REGION Network 2: Error handling
         A     #IN_Reset_fault_Fkt;
         R     #Temp_IO_Fault.FLT_Motorprotection;
         R     #Temp_IO_Fault.FLT_Min_Level;
         R     #Temp_IO_Fault.FLT_WRN_C_Max;
         R     #Temp_IO_Fault.FLT_C_Max;
         R     #Temp_IO_Fault.FLT_Filter_HP;
         R     #Temp_IO_Fault.FLT_Filter_backflow;
         R     #Temp_IO_Fault.FLT_cable_break;
         R     #Temp_IO_Fault.FLT_P_Max;
   //-----
         A     #IN_MotorProtection;
         AN    #Temp_IO_Fault.FLT_Motorprotection;
         S     #Temp_IO_Fault.FLT_Motorprotection;
         S     #IO_NewFault;
   //-----
         AN    #IN_Min_Level;
         AN    #Temp_IO_Fault.FLT_Min_Level;
         S     #Temp_IO_Fault.FLT_Min_Level;
         S     #IO_NewFault;
   //-----
         A     #IN_C_OilCooling;
         A     #Temp_IO_Status.Switch_on_Motor;
         =     #Temp_IO_Status.Act_Oilcooling;
   //-----
         AN    #IN_C_Max;
         AN    #Temp_IO_Fault.FLT_WRN_C_Max;
         S     #Temp_IO_Fault.FLT_WRN_C_Max;
         S     #IO_NewFault;
   //-----
         A     #Temp_IO_Fault.FLT_WRN_C_Max;
         L     S5T#5M;
         SD    #IN_Temperatur_Timer;
         A     #IN_Temperatur_Timer;
         AN    #Temp_IO_Fault.FLT_C_Max;
         S     #Temp_IO_Fault.FLT_C_Max;
         S     #IO_NewFault;
   //-----
         A     #Temp_IO_Status.Startup_Motor_finished;
         AN    #IN_F_Filter_ReturnLine;
         L     #IN_Delay_FilterError;
         SD    #IN_Filter_Timer;
   //-----
         AN    #IN_F_Filter_FeedLine;
         AN    #Temp_IO_Fault.FLT_Filter_HP;
         S     #Temp_IO_Fault.FLT_Filter_HP;
         S     #IO_NewFault;
   //-----
         A     #IN_Filter_Timer;
         AN    #IN_F_Filter_ReturnLine;
         AN    #Temp_IO_Fault.FLT_Filter_backflow;
         S     #Temp_IO_Fault.FLT_Filter_backflow;
         S     #IO_NewFault;
   //-----
         AN    #IN_P_lowerlimit;
         AN    #IN_P_upperLimit;
         S     #Temp_IO_Fault.FLT_cable_break;
         S     #IO_NewFault;
   //-----
         O     #IN_PRequestCycle;
         ON    #Temp_IO_Status.Startup_Motor_finished;
         O     #Temp_IO_Status.Request_from_CP;
         JC    NoFP;
   //-----
         L     #IN_P_BuildUpTime;
         AN    #Temp_IO_Status.MH_Hyd_OK;
         JC    TIME;
         L     #IN_P_OperationTime;
   TIME: NOP   0;
         A     #IN_P_upperLimit;
         A     #Temp_IO_Status.Act_PressureBuildUp;
         SD    #IN_Hydraulictimer;
         A     #IN_Hydraulictimer;
         AN    #Temp_IO_Fault.FLT_P_Max;
         S     #Temp_IO_Fault.FLT_P_Max;
         S     #IO_NewFault;
   //-----
   NoFP: NOP   0;
   //-----
END_REGION

REGION Network 3: An actual fault exist
   //-----
         O     #Temp_IO_Fault.FLT_Min_Level;
         O     #Temp_IO_Fault.FLT_Motorprotection;
         O     #Temp_IO_Fault.FLT_C_Max;
         O     #Temp_IO_Fault.FLT_P_Max;
         O     #Temp_IO_Fault.FLT_cable_break;
         O     #Temp_IO_Fault.FLT_WRN_C_Max;
         O     #Temp_IO_Fault.FLT_Filter_HP;
         O     #Temp_IO_Fault.FLT_Filter_backflow;
         =     #Temp_IO_Status.Fault_Exist;
   //-----
         O     #Temp_IO_Fault.FLT_Min_Level;
         O     #Temp_IO_Fault.FLT_Motorprotection;
         O     #Temp_IO_Fault.FLT_C_Max;
         O     #Temp_IO_Fault.FLT_P_Max;
         O     #Temp_IO_Fault.FLT_cable_break;
         =     #Temp_IO_Status.FaultLevel_1;
         S     #IO_FaultLevel_1;
   //-----
         O     #Temp_IO_Fault.FLT_WRN_C_Max;
         =     #Temp_IO_Status.FaultLevel_2;
         S     #IO_FaultLevel_2;
   //-----
         O     #Temp_IO_Fault.FLT_Filter_HP;
         O     #Temp_IO_Fault.FLT_Filter_backflow;
         =     #Temp_IO_Status.FaultLevel_3;
         S     #IO_FaultLevel_3;
   //-----
END_REGION

REGION Network 4
   //-----
         L     #IN_SwitchOffTime;
         T     #Temp_Motor_ON;
   //-----
         CALL  T_CONV
         ( IN  := #Temp_Motor_ON,
           OUT := #Temp_Motor_ON_ms
         );
   //-----
         L     #Temp_Motor_ON_ms;
         L     0;
         ==I;
         =     #Temp_No_switch_OFF;
   //-----
         L     #Temp_Motor_ON_ms;
         L     60000;  // 60 sec
         <D;
         =     #Temp_DelayTimeZero;
   //-----
END_REGION

REGION Network 5
   //-----
         O     #IN_ShotStroke_by_Piston;
         ON    #IN_KK_Manager_active;
         A     #IN_PRequestCycle;
         ON    #IN_P_lowerlimit;
         O     #Temp_IO_Status.Request_from_CP;
         O     #Temp_IO_Status.Act_Oilcooling;
         A     #Temp_IO_Status.MH_Hyd_OK;
         ON    #Temp_IO_Status.MH_Hyd_OK;
         AN    #Temp_No_switch_OFF;
         AN    #Temp_DelayTimeZero;
         L     #IN_SwitchOffTime;
         SF    #IN_SwitchOFFTimer;
         A     #IN_SwitchOFFTimer;
         =     #Temp_Motor_ON_Auto;
   //-----
         AN    #IN_OPMode_Automatic;
         R     #IN_SwitchOFFTimer;
   //-----
         O     #Temp_No_switch_OFF;
         O     #Temp_DelayTimeZero;
         O     #Temp_IO_Fault.Spare14;
         S     #Temp_Motor_ON_Auto;
   //-----
END_REGION

REGION Network 6: Request hydraulic
         O     #Temp_IO_Fault.FLT_Motorprotection;
         O     #Temp_IO_Fault.FLT_Min_Level;
         O     #Temp_IO_Fault.FLT_C_Max;
         O     #Temp_IO_Fault.FLT_cable_break;
         O     #Temp_IO_Fault.FLT_P_Max;
         =     #Temp_Fault_Hyd;
   //
         AN    #IN_Pos_of_Pause_ok;
         A     #IN_KK_Manager_active;
         ON    #IN_PauseTime;
         A     #Temp_IO_Status.Switch_Hydraulic_ON_OFF;
         A     #IN_OPMode_Manual;
         O     #IN_OPMode_Automatic;
         AN    #Temp_Fault_Hyd;
         AN    #IN_Fault_from_Extern;
         =     #Temp_IO_Status.Switch_on_Motor;
   //-
         A     #Temp_Motor_ON_Auto;
         A     #IN_OPMode_Automatic;
         O     #IN_OPMode_Manual;
         A     #Temp_IO_Status.Switch_on_Motor;
         =     #Temp_Switch_Motor_ON;
END_REGION

REGION Network 7: Motor control
         A     #Temp_IO_Status.Startup_Motor_finished;
         JC    NoM;
   //
         A     #Temp_Switch_Motor_ON;
         AN    #Temp_IO_Status.Act_Star;
         AN    #IN_Hydraulictimer;
         S     #Temp_IO_Status.Act_Main;
         S     #Temp_IO_Status.Act_Star;
         L     #IN_Star_Delta_Timer;
         SE    #IN_Hydraulictimer;
   //
         A     #Temp_Switch_Motor_ON;
         A     #Temp_IO_Status.Act_Star;
         AN    #IN_Hydraulictimer;
         S     #Temp_IO_Status.Startup_Motor_finished;
         R     #IN_Hydraulictimer;
   //
         A     #Temp_IO_Status.Startup_Motor_finished;
         AN    #Temp_IO_Status.MH_Hyd_OK;
         S     #Temp_IO_Status.Act_PressureBuildUp;
   //
   NoM:  NOP   0;
         AN    #Temp_Switch_Motor_ON;
         R     #Temp_IO_Status.Startup_Motor_finished;
         R     #Temp_IO_Status.Act_Main;
         R     #Temp_IO_Status.Act_Star;
         R     #Temp_IO_Status.Act_Delta;
   //
         AN    #Temp_IO_Status.Switch_on_Motor;
         R     #Temp_IO_Status.MH_Hyd_OK;
         R     #Temp_IO_Status.Act_PressureBuildUp;
END_REGION

REGION Network 8: Pressure valve control
   // Das Druckaufbauventil für die MK- Hydraulik wird angesteuert:
   // - Nachdem die Hydaulik angefordert wird (BA Auto oder Hydraulik EIN)
   // - Bei Anforderung aus dem Zyklusbaustein (3 Sekunden vor Ende der KLZ1 und
   //   der Schuß läuft), wenn es sich um eine Kolbenmaschine handelt muß der
   //   Schußhub laufen bei einer Pumpenmaschine sofort.
   // - Bei Anforderung aus dem Reinigungsbausteinen für die dauer von x Sekunden
         AN    #IN_P_upperLimit;
         A     #Temp_IO_Status.Act_PressureBuildUp;
         S     #Temp_IO_Status.MH_Hyd_OK;
         R     #Temp_IO_Status.Act_PressureBuildUp;
   //
         O     #IN_ShotStroke_by_Piston;
         ON    #IN_KK_Manager_active;
         A     #IN_PRequestCycle;
         AN    #IN_Option2SetPoints;
         ON    #IN_P_lowerlimit;
         O     #Temp_IO_Status.Request_from_CP;
         A     #Temp_IO_Status.Startup_Motor_finished;
         A     #Temp_IO_Status.MH_Hyd_OK;
         S     #Temp_IO_Status.Act_PressureBuildUp;
   //
         A     #Temp_IO_Status.MH_Hyd_OK;
         A     #Temp_IO_Status.Request_from_CP;
         A     #Temp_IO_Status.Startup_Motor_finished;
         JCN   NoRK;
   //
         SET;
         L     #IN_P_ClPistonTime;
         SE    #IN_Hydraulictimer;
   //
         AN    #IN_Hydraulictimer;
         R     #Temp_IO_Status.Request_from_CP;
         R     #IN_Hydraulictimer;
   //
   NoRK: NOP   0;
END_REGION

REGION Network 9: Outputs
   // Die hier praktizierte Art der Ansteuerung hat den Vorteil, dass die Parameter 
   // extern mit Dummys belegt werden können, wenn sie nicht gebraucht werden.
         A     #Temp_IO_Status.Act_PressureBuildUp;
         =     #OUT_PressureValve;
         A     #Temp_IO_Status.Act_Main;
         =     #OUT_Motor_MainsContactor;
         A     #Temp_IO_Status.Act_Star;
         =     #OUT_Motor_Star;
         A     #Temp_IO_Status.Act_Delta;
         =     #OUT_Motor_Delta;
         A     #Temp_IO_Status.Act_Oilcooling;
         =     #OUT_V_OilCooling;
         A     #Temp_IO_Status.MH_Hyd_OK;
         =     #OUT_Hydraulic_active;
END_REGION

REGION Network 10: State of drive: 1-> ON; 2-> Faulty; 3->Selected but not ON
         A     #Temp_IO_Status.MH_Hyd_OK;
         L     1;
         JC    tran;
   //-
         A     #Temp_IO_Status.Fault_Exist;
         L     2;
         JC    tran;
   //-
         A     #Temp_IO_Status.Switch_Hydraulic_ON_OFF;
         AN    #Temp_IO_Status.MH_Hyd_OK;
         L     3;
         JC    tran;
   //-
         L     0;
   tran: T     #Temp_IO_Status.State_Hydraulic;
END_REGION

REGION Network 11: Save data
   //-----
         CALL  BLKMOV
         ( SRCBLK  := #Temp_IO_Status,
           RET_VAL := #ERROR_CODE,
           DSTBLK  := #Anyzeiger1
         );
   //-----
         CALL  BLKMOV
         ( SRCBLK  := #Temp_IO_Fault,
           RET_VAL := #ERROR_CODE,
           DSTBLK  := #Anyzeiger2
         );
   //-----
END_REGION
END_FUNCTION

FUNCTION "FC025_Oszilloskop" : Void   // FC25, SCL
{ S7_Optimized_Access := 'FALSE' }
VERSION : 0.1
   VAR_TEMP
      i : Int;
      Baugruppe : Int;
      Index : Int;
      Wert : Int;
      connection : Int;
   END_VAR
BEGIN
   FOR #i := 1 TO 8 DO

     CASE "DB025_Oszilloskop".Graph[#i].Auswahl OF
       10:  CASE "DB025_Oszilloskop".Graph[#i].Komponente OF // Adresse
             20:  CASE "DB025_Oszilloskop".Graph[#i].Sensor OF  // Datenbaustein
                 101: "DB025_Oszilloskop".Graph[#i].Wert :=        // Bool
                     INT_TO_REAL(BOOL_TO_INT( PEEK_BOOL(area:=16#84,dbNumber:=WORD_TO_UINT("DB025_Oszilloskop".Graph[#i].DB_Nummer),byteOffset:="DB025_Oszilloskop".Graph[#i].Adresse,bitOffset:="DB025_Oszilloskop".Graph[#i].Bit) ) ) * "DB025_Oszilloskop".Graph[#i].Skalierung;  
                 102: "DB025_Oszilloskop".Graph[#i].Wert :=        // Byte
                     INT_TO_REAL( PEEK_BYTE(area:=16#84,dbNumber:=WORD_TO_UINT("DB025_Oszilloskop".Graph[#i].DB_Nummer),byteOffset:="DB025_Oszilloskop".Graph[#i].Adresse) ) * "DB025_Oszilloskop".Graph[#i].Skalierung; 
                 103: "DB025_Oszilloskop".Graph[#i].Wert :=        // Int
                     INT_TO_REAL( PEEK_WORD(area:=16#84,dbNumber:=WORD_TO_UINT("DB025_Oszilloskop".Graph[#i].DB_Nummer),byteOffset:="DB025_Oszilloskop".Graph[#i].Adresse) ) * "DB025_Oszilloskop".Graph[#i].Skalierung; 
                 104: "DB025_Oszilloskop".Graph[#i].Wert :=        // Dint
                     DINT_TO_REAL( PEEK_DWORD(area:=16#84,dbNumber:=WORD_TO_UINT("DB025_Oszilloskop".Graph[#i].DB_Nummer),byteOffset:="DB025_Oszilloskop".Graph[#i].Adresse) ) * "DB025_Oszilloskop".Graph[#i].Skalierung; 
                 105: "DB025_Oszilloskop".Graph[#i].Wert :=        // Real
                     DINT_TO_REAL( PEEK_DWORD(area:=16#84,dbNumber:=WORD_TO_UINT("DB025_Oszilloskop".Graph[#i].DB_Nummer),byteOffset:="DB025_Oszilloskop".Graph[#i].Adresse) ) * "DB025_Oszilloskop".Graph[#i].Skalierung; 
                 106: "DB025_Oszilloskop".Graph[#i].Wert :=        // Timer
                     REAL#0.0; 
               ELSE
                 "DB025_Oszilloskop".Graph[#i].Wert :=  REAL#0.0;
               END_CASE;
             21:  CASE "DB025_Oszilloskop".Graph[#i].Sensor OF  // Eingang
                 101: "DB025_Oszilloskop".Graph[#i].Wert :=        // Bool
                     INT_TO_REAL(BOOL_TO_INT( PEEK_BOOL(area:=16#81,dbNumber:=0,byteOffset:="DB025_Oszilloskop".Graph[#i].Adresse,bitOffset:="DB025_Oszilloskop".Graph[#i].Bit) ) ) * "DB025_Oszilloskop".Graph[#i].Skalierung;
                 102: "DB025_Oszilloskop".Graph[#i].Wert :=        // Byte
                     INT_TO_REAL( PEEK_BYTE(area:=16#81,dbNumber:=0,byteOffset:="DB025_Oszilloskop".Graph[#i].Adresse) ) * "DB025_Oszilloskop".Graph[#i].Skalierung; 
                 103: "DB025_Oszilloskop".Graph[#i].Wert :=        // Int
                     INT_TO_REAL( PEEK_WORD(area:=16#81,dbNumber:=0,byteOffset:="DB025_Oszilloskop".Graph[#i].Adresse) ) * "DB025_Oszilloskop".Graph[#i].Skalierung; 
                 104: "DB025_Oszilloskop".Graph[#i].Wert :=        // Dint
                     DINT_TO_REAL( PEEK_DWORD(area:=16#81,dbNumber:=0,byteOffset:="DB025_Oszilloskop".Graph[#i].Adresse) ) * "DB025_Oszilloskop".Graph[#i].Skalierung; 
                 105: "DB025_Oszilloskop".Graph[#i].Wert :=        // Real
                     REAL#0.0 ; 
               ELSE
                 "DB025_Oszilloskop".Graph[#i].Wert :=  REAL#0.0;
               END_CASE;
             22:  CASE "DB025_Oszilloskop".Graph[#i].Sensor OF  // Ausgang
                 101: "DB025_Oszilloskop".Graph[#i].Wert :=        // Bool
                     INT_TO_REAL(BOOL_TO_INT( PEEK_BOOL(area:=16#82,dbNumber:=0,byteOffset:="DB025_Oszilloskop".Graph[#i].Adresse,bitOffset:="DB025_Oszilloskop".Graph[#i].Bit) ) ) * "DB025_Oszilloskop".Graph[#i].Skalierung;
                 102: "DB025_Oszilloskop".Graph[#i].Wert :=        // Byte
                     INT_TO_REAL( PEEK_BYTE(area:=16#82,dbNumber:=0,byteOffset:="DB025_Oszilloskop".Graph[#i].Adresse) ) * "DB025_Oszilloskop".Graph[#i].Skalierung; 
                 103: "DB025_Oszilloskop".Graph[#i].Wert :=        // Int
                     INT_TO_REAL( PEEK_WORD(area:=16#82,dbNumber:=0,byteOffset:="DB025_Oszilloskop".Graph[#i].Adresse) ) * "DB025_Oszilloskop".Graph[#i].Skalierung; 
                 104: "DB025_Oszilloskop".Graph[#i].Wert :=        // Dint
                     DINT_TO_REAL( PEEK_DWORD(area:=16#82,dbNumber:=0,byteOffset:="DB025_Oszilloskop".Graph[#i].Adresse) ) * "DB025_Oszilloskop".Graph[#i].Skalierung; 
                 105: "DB025_Oszilloskop".Graph[#i].Wert :=        // Real
                     DINT_TO_REAL( PEEK_DWORD(area:=16#82,dbNumber:=0,byteOffset:="DB025_Oszilloskop".Graph[#i].Adresse) ) * "DB025_Oszilloskop".Graph[#i].Skalierung; 
               ELSE
                 "DB025_Oszilloskop".Graph[#i].Wert :=  REAL#0.0;
               END_CASE;
             23:  CASE "DB025_Oszilloskop".Graph[#i].Sensor OF  // Merker
                 101: "DB025_Oszilloskop".Graph[#i].Wert :=       // Bool
                     INT_TO_REAL(BOOL_TO_INT( PEEK_BOOL(area:=16#83,dbNumber:=0,byteOffset:="DB025_Oszilloskop".Graph[#i].Adresse,bitOffset:="DB025_Oszilloskop".Graph[#i].Bit) ) ) * "DB025_Oszilloskop".Graph[#i].Skalierung;
                 102: "DB025_Oszilloskop".Graph[#i].Wert :=        // Byte
                     INT_TO_REAL( PEEK_BYTE(area:=16#83,dbNumber:=0,byteOffset:="DB025_Oszilloskop".Graph[#i].Adresse) ) * "DB025_Oszilloskop".Graph[#i].Skalierung; 
                 103: "DB025_Oszilloskop".Graph[#i].Wert :=        // Int
                     INT_TO_REAL( PEEK_WORD(area:=16#83,dbNumber:=0,byteOffset:="DB025_Oszilloskop".Graph[#i].Adresse) ) * "DB025_Oszilloskop".Graph[#i].Skalierung; 
                 104: "DB025_Oszilloskop".Graph[#i].Wert :=        // Dint
                     DINT_TO_REAL( PEEK_DWORD(area:=16#83,dbNumber:=0,byteOffset:="DB025_Oszilloskop".Graph[#i].Adresse) ) * "DB025_Oszilloskop".Graph[#i].Skalierung; 
                 105: "DB025_Oszilloskop".Graph[#i].Wert :=         // Real
                     DINT_TO_REAL( PEEK_DWORD(area:=16#83,dbNumber:=0,byteOffset:="DB025_Oszilloskop".Graph[#i].Adresse) ) * "DB025_Oszilloskop".Graph[#i].Skalierung; ; 
               ELSE
                 "DB025_Oszilloskop".Graph[#i].Wert :=  REAL#0.0;
               END_CASE;
             24:  CASE "DB025_Oszilloskop".Graph[#i].Sensor OF  // Timer
                 106: "DB025_Oszilloskop".Graph[#i].Wert := REAL#0.0 ; // Timer
               ELSE
                 "DB025_Oszilloskop".Graph[#i].Wert :=  REAL#0.0;
               END_CASE;
           ELSE
             "DB025_Oszilloskop".Graph[#i].Wert :=  REAL#0.0;
           END_CASE;
       40:  CASE "DB025_Oszilloskop".Graph[#i].Sensor OF       // Behälter
             1:  "DB025_Oszilloskop".Graph[#i].Wert :=         // Durchfluss
                 REAL#0.0;               
             2:  "DB025_Oszilloskop".Graph[#i].Wert :=         // Druck
                 "DB602_PV_Tank".Tank["DB025_Oszilloskop".Graph[#i].Komponente].Pressure.PV_ActV.Value   * "DB025_Oszilloskop".Graph[#i].Skalierung;    
             3:  "DB025_Oszilloskop".Graph[#i].Wert :=         // Füllstand
                 "DB602_PV_Tank".Tank["DB025_Oszilloskop".Graph[#i].Komponente].Level.PV_ActV.Value      * "DB025_Oszilloskop".Graph[#i].Skalierung;         
             4:  "DB025_Oszilloskop".Graph[#i].Wert :=         // Gasbeladung
                 "DB602_PV_Tank".Tank["DB025_Oszilloskop".Graph[#i].Komponente].Nucleation.PV_ActV.Value * "DB025_Oszilloskop".Graph[#i].Skalierung;  
             5:  "DB025_Oszilloskop".Graph[#i].Wert :=         // Mischungsverhältnis         
                 REAL#40.0;              
             6:  "DB025_Oszilloskop".Graph[#i].Wert :=         // Temperatur
                 "DB602_PV_Tank".Tank["DB025_Oszilloskop".Graph[#i].Komponente].Temp.PV_ActV.Value       * "DB025_Oszilloskop".Graph[#i].Skalierung;        
           ELSE
             "DB025_Oszilloskop".Graph[#i].Wert :=  REAL#0.0;
           END_CASE;
        30:  CASE "DB025_Oszilloskop".Graph[#i].Sensor OF      // Pumpe
             1:  "DB025_Oszilloskop".Graph[#i].Wert :=         // Durchfluss
                 "DB608_PV_Metering".Metering["DB025_Oszilloskop".Graph[#i].Komponente].Flow.PV_ActV.Value *"DB025_Oszilloskop".Graph[#i].Skalierung;       
             2:  "DB025_Oszilloskop".Graph[#i].Wert :=         // Druck
                 "DB608_PV_Metering".Metering["DB025_Oszilloskop".Graph[#i].Komponente].Pressure.PV_ActV.Value  * "DB025_Oszilloskop".Graph[#i].Skalierung;    
             3:  "DB025_Oszilloskop".Graph[#i].Wert :=         // Füllstand
                 REAL#0.0;   
             4:  "DB025_Oszilloskop".Graph[#i].Wert :=         // Gasbeladung
                 REAL#0.0; 
             5:  "DB025_Oszilloskop".Graph[#i].Wert :=         // Mischungsverhältnis
                 "DB608_PV_Metering".Metering["DB025_Oszilloskop".Graph[#i].Komponente].MixingRatio.PV_ActV.Value  * "DB025_Oszilloskop".Graph[#i].Skalierung; 
             6:  "DB025_Oszilloskop".Graph[#i].Wert :=         // Temperatur
                 "DB608_PV_Metering".Metering["DB025_Oszilloskop".Graph[#i].Komponente].Temperature.PV_ActV.Value  * "DB025_Oszilloskop".Graph[#i].Skalierung; 
           ELSE
             "DB025_Oszilloskop".Graph[#i].Wert :=  REAL#0.0;
           END_CASE;
        20: #connection := 0;
                IF "DB025_Oszilloskop".Graph[#i].Komponente = "DB704_MH_Value".Mixinghead["DB025_Oszilloskop".Graph[#i].Nummer].MH_Connection[1].Pump_No THEN #connection := 1;  
                ELSIF "DB025_Oszilloskop".Graph[#i].Komponente = "DB704_MH_Value".Mixinghead["DB025_Oszilloskop".Graph[#i].Nummer].MH_Connection[2].Pump_No THEN #connection := 2;  
                ELSIF "DB025_Oszilloskop".Graph[#i].Komponente = "DB704_MH_Value".Mixinghead["DB025_Oszilloskop".Graph[#i].Nummer].MH_Connection[3].Pump_No THEN #connection := 3;  
                ELSIF "DB025_Oszilloskop".Graph[#i].Komponente = "DB704_MH_Value".Mixinghead["DB025_Oszilloskop".Graph[#i].Nummer].MH_Connection[4].Pump_No THEN #connection := 4;  
                ELSIF "DB025_Oszilloskop".Graph[#i].Komponente = "DB704_MH_Value".Mixinghead["DB025_Oszilloskop".Graph[#i].Nummer].MH_Connection[5].Pump_No THEN #connection := 5;  
                ELSIF "DB025_Oszilloskop".Graph[#i].Komponente = "DB704_MH_Value".Mixinghead["DB025_Oszilloskop".Graph[#i].Nummer].MH_Connection[6].Pump_No THEN #connection := 6;
                ELSE #connection := 0;
                END_IF;

           CASE "DB025_Oszilloskop".Graph[#i].Sensor OF        // Mischkopf    
             1:  "DB025_Oszilloskop".Graph[#i].Wert :=         // Durchfluss
                 REAL#0.0;             
             2:  "DB025_Oszilloskop".Graph[#i].Wert :=         // Druck
                 "DB604_PV_Mixinghead".Mixinghead["DB025_Oszilloskop".Graph[#i].Nummer].Pressure_Connection[#connection].PV_ActV.Value * "DB025_Oszilloskop".Graph[#i].Skalierung;  
             3:  "DB025_Oszilloskop".Graph[#i].Wert :=         // Füllstand
                 REAL#0.0;               
             4:  "DB025_Oszilloskop".Graph[#i].Wert :=         // Gasbeladung
                 REAL#0.0;             
             5:  "DB025_Oszilloskop".Graph[#i].Wert :=         // Mischungsverhältnis
                 REAL#0.0;                     
             6:  "DB025_Oszilloskop".Graph[#i].Wert :=         // Temperatur
                 "DB604_PV_Mixinghead".Mixinghead["DB025_Oszilloskop".Graph[#i].Nummer].Temperature_Connection[#connection].PV_ActV.Value * "DB025_Oszilloskop".Graph[#i].Skalierung;    
           ELSE
             "DB025_Oszilloskop".Graph[#i].Wert :=  REAL#0.0;
           END_CASE;
     ELSE
       "DB025_Oszilloskop".Graph[#i].Wert :=  REAL#0.0;
     END_CASE;
   END_FOR;
END_FUNCTION

FUNCTION "FC041_SwitchOverUnit" : Void   // FC41, STL
TITLE = Control of switch over units
{ S7_Optimized_Access := 'FALSE' }
AUTHOR : KT242
FAMILY : RS_KK
NAME : SWU
VERSION : 1.3
   VAR_INPUT
      IN_select_piston : Bool;   // Differentiation if programmblock is used by pump- or piston metering
      IN_filling_piston : Bool;   // Component piston in filling mode, used to switchover after strokes
      IN_OperationMode_valid : Bool;   // Operation mode valid
      IN_AcknoldgeFaults : Bool;   // Quit faults
      IN_cycle_running : Bool;   // During cycle is running no. of SWO is set by foaming program
      IN_PistonService : Bool;   // Piston service is selected to activate a switch over unit
      IN_Circulation_active : Bool;   // During active recirculation SWU will be switched over after a setted time
      IN_Circulation_HP_active : Bool;   // At high pressure circulation mixinghead no. is set by selected mixinghead
      IN_MH_No_at_FoamingCycle : Byte;   // Mixinghead number from foaming program to select SWU
      IN_MH_No_at_HP_Cycle : DWord;   // Mixinghead number from program block "operation mode" to select SWU by HP
      IN_StokeCounter : Counter;   // Counter of piston strokes to switch over to MH at piston machine
      IN_Amount_Strokes : Int;   // Setting of piston strokes to switch over to MH at piston machine
      IN_FlushingTimer : Timer;   // Timer flushing components between the mixingheads
      IN_SWU_FlushingTime : S5Time;   // Flushing time at each mixinghead at recirculation -> switchover to next MH
      IN_SwitchOverTimer : Timer;   // Timer to switch off and over between SWU's -> two SWU selected
      IN_SwitchOffTime : S5Time;   // Timevalue of increased activation of SWU at switch off
      IN_SwitchOverTime : S5Time;   // Timevalue of common activation of two SWU's during switch over
   END_VAR
   VAR_IN_OUT
      IO_Status : ANY;   // Speichern der Umschalteinheiten (USE)- Zustände für das Programm
      IO_Fault : ANY;
      IO_NewFault : Bool;
      IO_FaultLevel_1 : Bool;
      IO_FaultLevel_2 : Bool;
      IO_FaultLevel_3 : Bool;
   END_VAR
   VAR_TEMP
      Temp_IO_Status : "UDT041_SWU_State";
      TEMP_IO_Fault : "UDT1841_FLT_SWU";
      ERROR_CODE : Int;   // Error state of systemfunction "BLKMOV" Blockmove
      Anyzeiger1 : ANY;   // Pointer to copy thr array "IO_Status" and "Temp_IO_Status"
      Anyzeiger2 : ANY;   // Pointer to copy thr array "IO_Status" and "Temp_IO_Status"
      Baustein_Nr : Int;   // Merker zur Erkennung des Speicherbereiches der Bits "IO_Ziel_USE"
      Adresse_im_Baustein : DWord;   // and the start adress within the program block
      Freigaben_lokal : DWord;   // Intermidiate flags of release of switch over units (from UDT to DWORD)
      USE_Ventile_lokal : DWord;   // Zwischenspeicher der angesteuerten Umschalteinheiten (von UDT auf DWORD)
      Angef_USE_Nummer_lokal : DWord;   // Zwischenspeicher der angeforderten Umschalteinheiten (von UDT auf DWORD)
      Ziel_USE_lokal : DWord;   // Zwischenspeicher der auzusteuernden Umschalteinheiten (von UDT auf DWORD)
      U_A_Zeitwert : S5Time;   // Zeitwert bei der Unterscheidung ob eine USE um- oder abgeschaltet werden soll
      Temp_SWU_FlushingTime : S5Time;   // Zeitwert für die Spülzeit mindestens 3 Sekunden
      Spuelzeit_laeuft : Bool;   // Die Spülzeit der einzelnen Mischköpfe (USE) läuft und wird durchgetaktet
      Abschaltzeit_laeuft : Bool;   // Die Abschaltzeit der offenen USE läuft -> keine weitere USE angefordert
      Wiedereinschaltung : Bool;   // Es wurde innerhalb der Abschaltzeit Kreislauf etc. angeschaltet
   END_VAR
BEGIN

REGION Network 1: Saved data integration
   // Änderungen:
   // -------------------------------------------------------------------------------
   // Durch die Verwendung von + -1 bei der Ermittlung der angeforderten USE während 
   // des Zyklusses (Netzwerk 5) sind nur bis zu 16 Mischköpfe ansteuerbar.
   // Durch das umsetzen in Doppelworte (L     DW#16#1) wird eine Ansteuerung bis zu 
   // 32 Mischköpfe möglich
   // 
   // v.d.Geest       19.01.2005
   // -------------------------------------------------------------------------------
   // Wenn im Rechner ein Mischkopf als folgender Teilschuß angewählt wurde, dessen 
   // USE aber nicht freigegeben war kam es zu einer Max. Druck- Störung.
   // Um dieses zu vermeiden wurde eine neue Störung "USE_nicht_freigegeben" im 
   // Netzwerk 7 ab Zeile 49 eingebunden.
   // 
   // v.d.Geest       27.10.2003
   // -------------------------------------------------------------------------------
   // Die Ansteuerung der "Um_Abschaltzeit" funktionierte so nicht:
   // Bei Anwahl Kreislauf aus dem Stillstand lief die "Um_Abschaltzeit" ab, obwohl 
   // vorher kein weiterer Mischkopf angewählt wurde. 
   // Ebenso wurde die gesamte Abschaltzeit abgewartet wenn zwischen dem Auschalten 
   // des Kreislaufes über zB. MK01 und dem winschalten des Kreislaufes über zB. MK02 
   // weniger als 5 Sekunden (Abschaltzeit) lagen.
   // Die Auswirkungen waren zu spüren der Anwahl des HD- Kreislaufes, da dieser erst 
   // gestartet wurde wenn die "Um_Abschaltzeit" abgelaufen war.
   // Das alte Bit "Um_Abschaltzeit" im UDT wurde in "Umschaltzeit" (wichtig bei 
   // schnellem Druckaufbau und bei Ansteuerung des Reinigungskolbens) umbenannt und 
   // ein neues Bit "Abschaltzeit" wurde erstellt.
   // Bei Übernahme bitte UDT 41 mit einspielen.
   // 
   // v.d.Geest       11.04.2003
   // -------------------------------------------------------------------------------
         LAR1;
         L;
         LAR2;
   //
         L     W[AR2, P#0.0];  // Bytes
         T     W[AR1, P#0.0];
         L     W [ AR2 , P#2.0 ];  // Amount of bytes
         T     W[AR1, P#2.0];
         L     W [ AR2 , P#4.0 ];  // Block no,
         T     W[AR1, P#4.0];
         L     D [ AR2 , P#6.0 ];  // Startadress of datas
         T     D[AR1, P#6.0];
   //
         CALL  BLKMOV
         ( SRCBLK  := #Anyzeiger1,
           RET_VAL := #ERROR_CODE,
           DSTBLK  := #Temp_IO_Status
         );

         LAR1;
         L;
         LAR2;
   //
         L     W[AR2, P#0.0];  // Bytes
         T     W[AR1, P#0.0];
         L     W [ AR2 , P#2.0 ];  // Amount of bytes
         T     W[AR1, P#2.0];
         L     W [ AR2 , P#4.0 ];  // Block no,
         T     W[AR1, P#4.0];
         L     D [ AR2 , P#6.0 ];  // Startadress of datas
         T     D[AR1, P#6.0];
   //
         CALL  BLKMOV
         ( SRCBLK  := #Anyzeiger2,
           RET_VAL := #ERROR_CODE,
           DSTBLK  := #TEMP_IO_Fault
         );
   //
END_REGION

REGION Network 2: Störungen quittieren
         A     #IN_AcknoldgeFaults;
         R     #TEMP_IO_Fault.FLT_open_SWU_disabelt;
         R     #TEMP_IO_Fault.FLT_No_SWU_selected;
         R     #TEMP_IO_Fault.FLT_Sel_SWU_not_released;
END_REGION

REGION Network 3: Datenschieben
   //_______________________________________________________________
   // Schieben der USE- Freigaben auf lokalen DWord- Bereich
   //
         L;
         LAR2;
         L;
         LAR1;
   //
         L     LD [ AR2 , P#8.0 ];
         T     LD[AR1, P#0.0];
   //_______________________________________________________________
   // Schieben der Ziel- USE vom Rechner auf lokalen DWord- Bereich
   //
         L;
         LAR2;
         L;
         LAR1;
   //
         L     LD [ AR2 , P#12.0 ];
         T     LD[AR1, P#0.0];
   //_______________________________________________________________
   // Schieben der offenen USE auf lokalen DWord- Bereich
   //
         L;
         LAR1;
   //
         L     LD [ AR2 , P#16.0 ];
         T     LD[AR1, P#0.0];
END_REGION

REGION Network 4: Allgemein Verwaltung der angeforderten USE
         L     #Freigaben_lokal;
         L     0;
         <>D;
         =     #Temp_IO_Status.Min_1_SWU_release;
   //
         L     #USE_Ventile_lokal;
         L     #Freigaben_lokal;
         AD;
         <>D;
         =     #Temp_IO_Status.Open_SWU_disabelt;
   //
         ON    #IN_cycle_running;
         R     #Temp_IO_Status.CycleStarted;
   //
         A     #IN_cycle_running;
         A(;
         L     #IN_MH_No_at_FoamingCycle;
         L     0;
         <>I;
         );
         O     #Temp_IO_Status.CycleStarted;
         JC    ZYKL;
   //
         A     #IN_Circulation_HP_active;
         JC    HD;
   //
         O     #IN_Circulation_active;
         O     #IN_PistonService;
         A     #Temp_IO_Status.Min_1_SWU_release;
         JC    KK;
END_REGION

REGION Network 5: Keine USE angefordert
         L     0;
         T     #Angef_USE_Nummer_lokal;
   //
         SET;
         R     #IN_StokeCounter;
         R     #Temp_IO_Status.Hubcounter_OK;
         R     #IN_FlushingTimer;
   //
         CLR;
         SP    #IN_FlushingTimer;
   //
         JU    N05A;
END_REGION

REGION Network 6: Zyklus läuft oder Kreislauf Hochdruck
   ZYKL: NOP   0;
         S     #Temp_IO_Status.CycleStarted;
   //-
         L     0;
         L     #IN_MH_No_at_FoamingCycle;
         ==I;
         JC    NoUS;
         L     16#0000_0001;
         -D;
         L     16#0000_0001;
         SLD;
         JU    Next;
   NoUS: L     #Ziel_USE_lokal;
   Next: T     #Angef_USE_Nummer_lokal;
         JU    N05A;
   //
   HD:   L     #IN_MH_No_at_HP_Cycle;
         T     #Angef_USE_Nummer_lokal;
         JU    N05A;
END_REGION

REGION Network 7: Unterscheidung RS oder KK für USE- Spülung
   KK:   AN    #IN_select_piston;
         JC    RS;
   //
         A     #IN_Circulation_active;
         A     #IN_filling_piston;
         CU    #IN_StokeCounter;
   //
         L     #IN_Amount_Strokes;
         LC    #IN_StokeCounter;
         ==I;
         R     #IN_StokeCounter;
         =     #Temp_IO_Status.Hubcounter_OK;
   //
   RS:   L     0;
         L     #Temp_IO_Status.SWU_for_Circulation;
         ==D;
         JC    ERST;
         JU    SPUE;
   ERST: L     1;
         T     #Temp_IO_Status.SWU_for_Circulation;
   //
   SPUE: L     #IN_SWU_FlushingTime;
         T     #Temp_SWU_FlushingTime;
         L     S5T#3S;
         >D;
         JC    STRT;
         T     #Temp_SWU_FlushingTime;
   //
   STRT: A(;
         AN    #IN_FlushingTimer;
         AN    #IN_select_piston;
         O;
         AN    #Temp_IO_Status.Hubcounter_OK;
         A     #IN_select_piston;
         );
         A(;
         L     #Temp_IO_Status.SWU_for_Circulation;
         L     #Freigaben_lokal;
         AD;
         ==D;
         );
         =     #Spuelzeit_laeuft;
   //
         A     #Spuelzeit_laeuft;
         AN    #IN_select_piston;
         L     #Temp_SWU_FlushingTime;
         SD    #IN_FlushingTimer;
   //
         A     #Spuelzeit_laeuft;
         JC    RED;
   //
   TAKT: L     #Temp_IO_Status.SWU_for_Circulation;
         SLD   1;
         JP    USE1;
         JU    TEST;
   //
   USE1: L     1;
   //
   TEST: T     #Temp_IO_Status.SWU_for_Circulation;
         L     #Freigaben_lokal;
         AD;
         <>D;
         JC    TAKT;
   //
   RED:  L     #Temp_IO_Status.SWU_for_Circulation;
         T     #Angef_USE_Nummer_lokal;
END_REGION

REGION Network 8: Abschaltzeit / Umschaltzeit / USE- Ansteuerung
   N05A: L     #Angef_USE_Nummer_lokal;
         L     0;
         ==D;
         =     #Abschaltzeit_laeuft;
         S     #Temp_IO_Status.Stoptime_runs;
   //
         AN    #Abschaltzeit_laeuft;
         A     #Temp_IO_Status.Stoptime_runs;
         =     #Wiedereinschaltung;
         R     #Temp_IO_Status.Stoptime_runs;
         JC    Cl_T;
   //
         L     #IN_SwitchOverTime;
         AN    #Abschaltzeit_laeuft;
         JC    Zeit;
         L     #IN_SwitchOffTime;
   Zeit: T     #U_A_Zeitwert;
   //
         A(;
         L     #Ziel_USE_lokal;  // USE_Ventile
         L     0;
         <>D;
         );
         A(;
         L     #Angef_USE_Nummer_lokal;
         L     #Ziel_USE_lokal;  // USE_Ventile
         <>D;
         );
         L     #U_A_Zeitwert;
         SE    #IN_SwitchOverTimer;
   //
         AN    #IN_SwitchOverTimer;
         R     #Temp_IO_Status.Stoptime_runs;
   //
         A     #IN_SwitchOverTimer;
         AN    #Temp_IO_Status.Stoptime_runs;
         =     #Temp_IO_Status.Switchingtime_runs;
         JU    ZUSE;
   //
   Cl_T: NOP   0;
         CLR;
         SP    #IN_SwitchOverTimer;
   //
   ZUSE: L     #Angef_USE_Nummer_lokal;
         L     #Freigaben_lokal;
         AD;
         T     #Ziel_USE_lokal;  // USE_Ventile
   //
         A(;
         L     #Angef_USE_Nummer_lokal;
         L     0;
         <>D;
         );
         A(;
         L     #Ziel_USE_lokal;  // USE_Ventile
         L     0;
         ==D;
         );
         =     #Temp_IO_Status.SWU_not_released;
   //_______________________________________________________________
   // Schieben der allein offenen USE auf den Status - Bereich
   //
         L;
         LAR2;
         L;  // USE_Ventile
         LAR1;
   //
         L     LD[AR1, P#0.0];  // USE_Ventile
         T     LD [ AR2 , P#20.0 ];  // Temp_Status.Offene_USE_allein
   //
         O     #Temp_IO_Status.Switchingtime_runs;
         O     #Temp_IO_Status.Stoptime_runs;
         JCN   OUSE;
   //
         L     #Ziel_USE_lokal;
         L     #USE_Ventile_lokal;
         OW;
         T     #USE_Ventile_lokal;
   //_______________________________________________________________
   // Ablöschen der allein offenen USE auf den Status - Bereich
   //
         L;
         LAR2;
   //
         L     0;
         T     LD [ AR2 , P#20.0 ];  // Temp_Status.Offene_USE_allein
   //
         JU    M017;
   //
   OUSE: NOP   0;
   //
         L     #Ziel_USE_lokal;
         T     #USE_Ventile_lokal;
   //
   M017: NOP   0;
   //
         L     #USE_Ventile_lokal;
         L     0;
         ==D;
         R     #Temp_IO_Status.SWU_OK;
         JC    NUSE;
   //
   M012: NOP   0;
         TAK;
         SRD   1;
         JZ    M012;
         ==I;
         =     #Temp_IO_Status.SWU_OK;
   //
   NUSE: NOP   0;
END_REGION

REGION Network 9
   //_______________________________________________________________
   // Schieben der offenen USE auf den "IO_Status"- Bereich
   //
         L;
         LAR2;
         L;
         LAR1;
   //
         L     LD[AR1, P#0.0];  // USE_Ventile
         T     LD [ AR2 , P#16.0 ];  // Temp_Status.Open_SWU
   //_______________________________________________________________
   // Schieben der lokalen Ziel- USE auf den Ziel- USE- Bereich
   //
         L;
         LAR2;
         L;
         LAR1;
         L     LD [ AR1 , P#0.0 ];  // Ziel_USE_Lokal
         T     LD [ AR2 , P#12.0 ];  // Temp_Status.Target_SWU
   //_______________________________________________________________
   //
END_REGION

REGION Network 10
         L     0;
         A     #Temp_IO_Status.Target_SWU."01";
         JCN   nMH01;
         +     1;
         JU    NoHMopen;
   nMH01:NOP   0;
         A     #Temp_IO_Status.Target_SWU."02";
         JCN   nMH02;
         +     2;
         JU    NoHMopen;
   nMH02:NOP   0;
         A     #Temp_IO_Status.Target_SWU."03";
         JCN   nMH03;
         +     3;
         JU    NoHMopen;
   nMH03:NOP   0;
         A     #Temp_IO_Status.Target_SWU."04";
         JCN   nMH04;
         +     4;
         JU    NoHMopen;
   nMH04:NOP   0;
         A     #Temp_IO_Status.Target_SWU."05";
         JCN   nMH05;
         +     5;
         JU    NoHMopen;
   nMH05:NOP   0;
         A     #Temp_IO_Status.Target_SWU."06";
         JCN   nMH06;
         +     6;
         JU    NoHMopen;
   nMH06:NOP   0;
         A     #Temp_IO_Status.Target_SWU."07";
         JCN   nMH07;
         +     7;
         JU    NoHMopen;
   nMH07:NOP   0;
         A     #Temp_IO_Status.Target_SWU."08";
         JCN   nMH08;
         +     8;
         JU    NoHMopen;
   nMH08:NOP   0;
         A     #Temp_IO_Status.Target_SWU."09";
         JCN   nMH09;
         +     9;
         JU    NoHMopen;
   nMH09:NOP   0;
         A     #Temp_IO_Status.Target_SWU."10";
         JCN   nMH10;
         +     10;
         JU    NoHMopen;
   nMH10:NOP   0;
         A     #Temp_IO_Status.Target_SWU."11";
         JCN   nMH11;
         +     11;
         JU    NoHMopen;
   nMH11:NOP   0;
         A     #Temp_IO_Status.Target_SWU."12";
         JCN   nMH12;
         +     12;
         JU    NoHMopen;
   nMH12:NOP   0;
         A     #Temp_IO_Status.Target_SWU."13";
         JCN   nMH13;
         +     13;
         JU    NoHMopen;
   nMH13:NOP   0;
         A     #Temp_IO_Status.Target_SWU."14";
         JCN   nMH14;
         +     14;
         JU    NoHMopen;
   nMH14:NOP   0;
         A     #Temp_IO_Status.Target_SWU."15";
         JCN   nMH15;
         +     15;
         JU    NoHMopen;
   nMH15:NOP   0;
         A     #Temp_IO_Status.Target_SWU."16";
         JCN   nMH16;
         +     16;
         JU    NoHMopen;
   nMH16:NOP   0;

   NoHMopen:NOP   0;
         T     #Temp_IO_Status.ActualSWU;
END_REGION

REGION Network 11: Error handling
         A     #Temp_IO_Status.Open_SWU_disabelt;
         AN    #TEMP_IO_Fault.FLT_open_SWU_disabelt;
         S     #TEMP_IO_Fault.FLT_open_SWU_disabelt;
         S     #IO_NewFault;
   //-----
         AN    #Temp_IO_Status.Min_1_SWU_release;
         A     #IN_OperationMode_valid;
         AN    #TEMP_IO_Fault.FLT_No_SWU_selected;
         S     #TEMP_IO_Fault.FLT_No_SWU_selected;
         S     #IO_NewFault;
   //-----
         A     #Temp_IO_Status.SWU_not_released;
         AN    #TEMP_IO_Fault.FLT_Sel_SWU_not_released;
         S     #TEMP_IO_Fault.FLT_Sel_SWU_not_released;
         S     #IO_NewFault;
   //-----
         O     #TEMP_IO_Fault.FLT_open_SWU_disabelt;
         O     #TEMP_IO_Fault.FLT_No_SWU_selected;
         O     #TEMP_IO_Fault.FLT_Sel_SWU_not_released;
         =     #Temp_IO_Status.FaultLevel_1;
         S     #IO_FaultLevel_1;
   //-----
         CLR;
         =     #Temp_IO_Status.FaultLevel_2;
         S     #IO_FaultLevel_2;
   //-----
         CLR;
         =     #Temp_IO_Status.FaultLevel_3;
         S     #IO_FaultLevel_3;
END_REGION

REGION Network 12: Save data
         CALL  BLKMOV
         ( SRCBLK  := #Temp_IO_Status,
           RET_VAL := #ERROR_CODE,
           DSTBLK  := #Anyzeiger1
         );
   //
         CALL  BLKMOV
         ( SRCBLK  := #TEMP_IO_Fault,
           RET_VAL := #ERROR_CODE,
           DSTBLK  := #Anyzeiger2
         );
   //
END_REGION
END_FUNCTION

FUNCTION "FC042_MixingHead" : Void   // FC42, STL
TITLE = Control of mixinghead valve
{ S7_Optimized_Access := 'FALSE' }
AUTHOR : KT242
FAMILY : RS_KK
NAME : MHead
VERSION : 1.1
   VAR_INPUT
      IN_SWU_openValve : "UDT001_DWord_1_32";
      IN_OPMode_Automatic : Bool;
      IN_OPMode_Production : Bool;
      IN_OPMode_Test : Bool;
      IN_Error_Level_1 : Bool;
      IN_SWU_OK : Bool;
      IN_Release_Foamingcycle : Bool;
      IN_ExternalRel_Foaming : Bool;
      IN_ToleranceOK_Foaming : Bool;
      IN_Foaming_Active : Bool;
   END_VAR
   VAR_IN_OUT
      IO_Status : ANY;
   END_VAR
   VAR_TEMP
      Temp_IO_Status : "UDT042_MH_Select";
      Temp_ERROR_CODE : Int;
      Anyzeiger : ANY;
      Temp_DataBlock_No : Int;
      Temp_AddressInDatablock : DWord;
      Temp_ReleaseMH : DWord;
      Temp_MHValve : DWord;
      Temp_Shotcounter : DWord;
      Temp_SWU_Valve : DWord;
      Temp_HF_Foaming_active : Bool;
   END_VAR
BEGIN

REGION Network 1: Saved data integration
         LAR1;
         L;
         LAR2;
   //
         L     W[AR2, P#0.0];  // Bytes
         T     W[AR1, P#0.0];
         L     W[AR2, P#2.0];  //Amount of bytes
         T     W[AR1, P#2.0];
         L     W[AR2, P#4.0];  //Block no,
         T     W[AR1, P#4.0];
         L     D[AR2, P#6.0];  //Startadress of datas
         T     D[AR1, P#6.0];
   //
         CALL  BLKMOV
         ( SRCBLK  := #Anyzeiger,
           RET_VAL := #Temp_ERROR_CODE,
           DSTBLK  := #Temp_IO_Status
         );
   //
END_REGION

REGION Network 2: Data shifting
   //_______________________________________________________________
   // Schieben der Offenen- USE auf lokalen DWord- Bereich
   //
         L;  //
         LAR1;  //
         L     W[AR1, P#0.0];  //
         T     #Temp_DataBlock_No;  //
   //
         L     D[AR1, P#2.0];
         T     #Temp_AddressInDatablock;  //
         LAR2;  //
         L;  //
         LAR1;  //
   //
         OPN   DB[ #Temp_DataBlock_No];  //
         L     DBD[AR2, P#0.0];  //
         T     LD[AR1, P#0.0];  //
   //_______________________________________________________________
   // Schieben der Freigegeben MK's auf lokalen DWord- Bereich
   //
         L;  //
         LAR2;  //
         L;  //
         LAR1;  //
   //
         L     LD[AR2, P#0.0];  //
         T     LD[AR1, P#0.0];  //
END_REGION

REGION Network 3: Mixingheadcontrol of 32 mixing heads
         L     #Temp_SWU_Valve;
         T     #Temp_MHValve;
   //
         A(;
         L     #Temp_ReleaseMH;
         L     #Temp_MHValve;
         AD;
         L     0;
         <>D;
         );
         A     #IN_OPMode_Automatic;
         A     #IN_Release_Foamingcycle;
         A     #IN_SWU_OK;
         AN    #IN_Error_Level_1;
         A     #IN_ExternalRel_Foaming;
         A     #Temp_IO_Status.Cleaningpiston_OK;
         A     #IN_ToleranceOK_Foaming;
         JC    ENDE;
   //
         L     0;
         T     #Temp_MHValve;
   ENDE: NOP   0;
END_REGION

REGION Network 4: Activate mechanical shotcounter
         A(;
         A     #IN_OPMode_Production;
         AN    #IN_OPMode_Test;
         A     #IN_Foaming_Active;
         JNB   _001;
   //
         L     #Temp_MHValve;
         T     #Temp_Shotcounter;
         SET;
   //
         SAVE;
         CLR;
   _001: A     BR;
         );
         =     #Temp_HF_Foaming_active;
   //
         A     #Temp_HF_Foaming_active;
         NOT;
         JNB   _002;
         L     0;
         T     #Temp_Shotcounter;
   _002: NOP   0;
END_REGION

REGION Network 5: Add up shot counter of the value 1 per 1 SPS- cycle
         A(;
         A(;
         A     #Temp_HF_Foaming_active;
         BLD   100;
         FP    #Temp_IO_Status.Counterrampe;
         =     #Temp_IO_Status.ImpCounterOn;
         );
         JNB   _003;
         L     1;
         T     #Temp_IO_Status.Countervalue;
         SET;
         SAVE;
         CLR;
   _003: A     BR;
         );
         NOT;
         JNB   _006;
         L     0;
         T     #Temp_IO_Status.Countervalue;
   _006: NOP   0;
END_REGION

REGION Network 6: Data transfer
   //_______________________________________________________________
   // Schieben der lokalen MK- Ventile auf den "IO_Status"- Bereich
   //
         L;  //
         LAR2;  //
         L;  //
         LAR1;  //
         L     LD[AR1, P#0.0];  //
         T     LD[AR2, P#4.0];  //
   //_______________________________________________________________
   // Schieben der lokalen Schußzähler auf den "IO_Status"- Bereich
   //
         L;  //
         LAR1;  //
         L     LD[AR1, P#0.0];  //
         T     LD[AR2, P#8.0];  //
END_REGION

REGION Network 7: Save data
         CALL  BLKMOV
         ( SRCBLK  := #Temp_IO_Status,
           RET_VAL := #Temp_ERROR_CODE,
           DSTBLK  := #Anyzeiger
         );
   //
END_REGION
END_FUNCTION

FUNCTION "FC051_ComponentGeneral" : Void   // FC51, SCL
{ S7_Optimized_Access := 'FALSE' }
VERSION : 0.1
   VAR_TEMP
      i : Int;
   END_VAR
BEGIN
   FOR #i := 1 TO 12 DO
     // Delete all Fault information at the Main Window
     "DB613_Komponent_State".GroupStatus[#i].FaultExist := 0;
   END_FOR;

   FOR #i := 1 TO "DB790_PlantParameter".AmountMeteringUnits DO
     "DB613_Komponent_State".GroupStatus[#i].ColorTankFlow :="DB702_Tank_Value".Tank["DB753_MeteringPump".Pump[#i].TankNo].Color;
     "DB613_Komponent_State".GroupStatus[#i].FaultExist := "DB613_Komponent_State".EdgeFilter[#i].FLT_Exist OR
                                                           "DB613_Komponent_State".FeedPump[#i].FLT_Exist OR
                                                           "DB613_Komponent_State".MeteringPump[#i].FLT_Exist OR
                                                           "DB613_Komponent_State".HeatexchangerHP[#i].Fault_Exist OR
                                                           "DB613_Komponent_State".HeatexchangerLP[#i].Fault_Exist OR
                                                           "DB823_Error_Metering".MeteringPump[#i].FLT_MotorFan;

       IF "DB753_MeteringPump".Pump[#i].WithFlowFactor = False THEN
           "DB753_MeteringPump".Pump[#i].FlowFactor := 1.00;
       END_IF;

   END_FOR;
END_FUNCTION

FUNCTION "FC053_MeteringPump" : Void   // FC53, STL
TITLE = Control of metering pumps 2 speeds or frequency units
{ S7_Optimized_Access := 'FALSE' }
AUTHOR : KT242
FAMILY : RS
NAME : PUMP